(* Logix 5000 project; controller FV vendor 1 type 14 code 217 rev 31.11; software revision 31.00; part 7 of 63 *)
(* tags used below, declared in another part *)
   CWD : CHECKWORD_FLAGS;
   Dummy : BOOL;
   FR_B240 : INT[255];   // DEBOUNCE Debounce Flags
   fr_chk_temp : DINT;
   FR_copy_how_many : DINT;
   FR_data_file_value_to_move : DINT;
   FR_from_data_file : DINT;
   FR_from_data_offset : DINT;
   FR_FV26_HLP01 : PlantItem;   // FV26_HLP01
   FR_FV26_LLP01 : PlantItem;   // FV26_LLP01
   FR_FV27_HLP01 : PlantItem;   // FV27_HLP01
   FR_FV27_LLP01 : PlantItem;   // FV27_LLP01
   FR_FV28_HLP01 : PlantItem;   // FV28_HLP01
   FR_FV28_LLP01 : PlantItem;   // FV28_LLP01
   FR_FV29_HLP01 : PlantItem;   // FV29_HLP01
   FR_FV29_LLP01 : PlantItem;   // FV29_LLP01
   FR_FV30_HLP01 : PlantItem;   // FV30_HLP01
   FR_FV30_LLP01 : PlantItem;   // FV30_LLP01
   FR_FV31_HLP01 : PlantItem;   // FV31_HLP01
   FR_N10 : INT[265];   // FV_AGING Comms to FV Aging PL C
   FR_N100 : INT[265];   // FV FILLING
   FR_N110 : INT[265];   // GREEN BEER Green Beer Main
   FR_N120 : INT[265];   // YEAST CROP Yeast Cropping Main
   FR_N13 : INT[265];   // MV_ROUTE Comms to MV Routing PLC
   FR_N130 : INT[265];   // FILTRATE Filtrate Return
   FR_N14 : INT[265];   // MVFV CIP Comms to MVFV CIP Un it PLC
   FR_N140 : INT[265];   // CIP
   FR_N142 : INT[265];   // CIP
   FR_N143 : INT[265];   // CIP
   FR_N150 : INT[265];   // Original N File From SLC, No Description Available
   FR_N160 : INT[265];   // VESSEL Vessel Working Direc tory
   FR_N170 : INT[265];   // Original N File From SLC, No Description Available
   FR_N180 : INT[265];   // Original N File From SLC, No Description Available
   FR_N198 : INT[265];   // Original N File From SLC, No Description Available
   FR_N20 : INT[265];   // GENERAL General Purpose Setp oints
   FR_N200 : INT[265];   // ANALOG_IN Analog Inputs
   FR_N201 : INT[265];   // Original N File From SLC, No Description Available
   FR_N207 : INT[265];   // Original N File From SLC, No Description Available
   FR_N21 : INT[265];   // CHASE_V FV Filling Beer Chas e Volumes
   FR_N210 : INT[265];   // ANALOG_OUT Analog Outputs
   FR_N220 : INT[265];   // CHECKLIST Checklist Loop Contr ollers
   FR_N225 : INT[265];   // Original N File From SLC, No Description Available
   FR_N226 : INT[265];   // Original N File From SLC, No Description Available
   FR_N245 : INT[265];   // CHECKWORD Checkword Loop Contr ol
   FR_N252 : INT[265];   // OUTPUT_PTR Checkword Pointers t o output flags in B2 50
   FR_N253 : INT[265];   // EN_POINT Pointers to energise d input flags in B25 1
   FR_N254 : INT[265];   // DEN_POINT Pointers to deenergi sed input flags in B 251
   FR_N255 : INT[265];   // CHECKWORDS
   FR_N26 : INT[265];   // FV26
   FR_N27 : INT[265];   // FV27
   FR_N28 : INT[265];   // FV28
   FR_N29 : INT[265];   // FV29
   FR_N30 : INT[265];   // FV30
   FR_N31 : INT[265];   // FV31
   FR_N36 : INT[265];   // Original N File From SLC, No Description Available
   FR_N37 : INT[265];   // Original N File From SLC, No Description Available
   FR_N46 : INT[265];   // Original N File From SLC, No Description Available
   FR_N47 : INT[265];   // Original N File From SLC, No Description Available
   FR_N7 : INT[265];   // INTEGER
   FR_N99 : INT[265];   // COMMENT Comment Lines
   FR_T242 : TIMER[255];   // DEBOUNCE
   FR_T243 : TIMER[255];   // DEBOUNCE
   FR_to_data_file : DINT;
   FR_to_data_offset : DINT;
(* FR_Common, continued *)

ROUTINE FR_CHECK_LIST_220   (* ladder *)
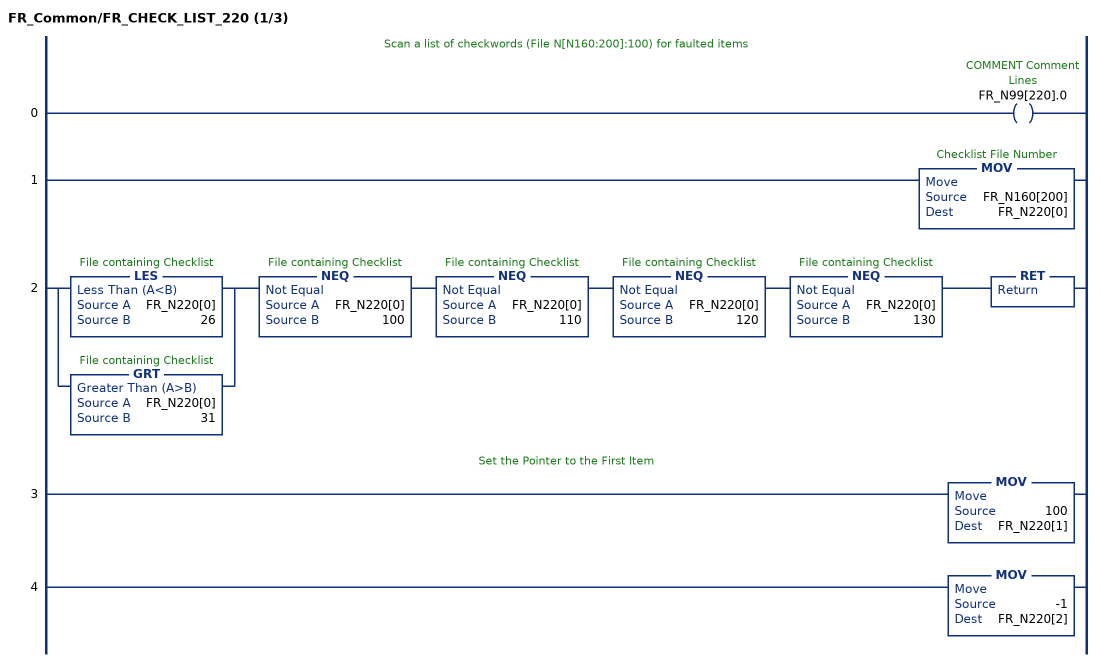
   // Scan a list of checkwords (File N[N160:200]:100) for faulted items
   0: OTE(FR_N99[220].0);
   1: MOV(FR_N160[200],FR_N220[0]);
   2: [LES(FR_N220[0],26) ,GRT(FR_N220[0],31) ]NEQ(FR_N220[0],100)NEQ(FR_N220[0],110)NEQ(FR_N220[0],120)NEQ(FR_N220[0],130)RET();
   // Set the Pointer to the First Item
   3: MOV(100,FR_N220[1]);
   4: MOV(-1,FR_N220[2]);
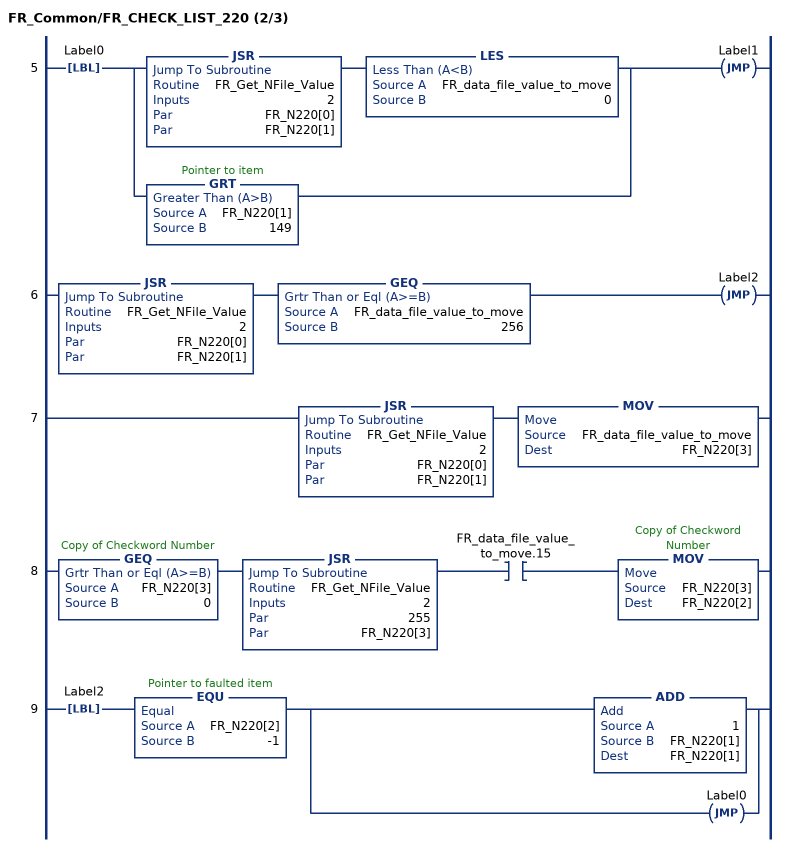
   5: LBL(Label0)[JSR(FR_Get_NFile_Value,2,FR_N220[0],FR_N220[1]) LES(FR_data_file_value_to_move,0) ,GRT(FR_N220[1],149) ]JMP(Label1);
   6: JSR(FR_Get_NFile_Value,2,FR_N220[0],FR_N220[1])GEQ(FR_data_file_value_to_move,256)JMP(Label2);
   7: JSR(FR_Get_NFile_Value,2,FR_N220[0],FR_N220[1])MOV(FR_data_file_value_to_move,FR_N220[3]);
   8: GEQ(FR_N220[3],0)JSR(FR_Get_NFile_Value,2,255,FR_N220[3])XIC(FR_data_file_value_to_move.15)MOV(FR_N220[3],FR_N220[2]);
   9: LBL(Label2)EQU(FR_N220[2],-1)[ADD(1,FR_N220[1],FR_N220[1]) ,JMP(Label0) ];
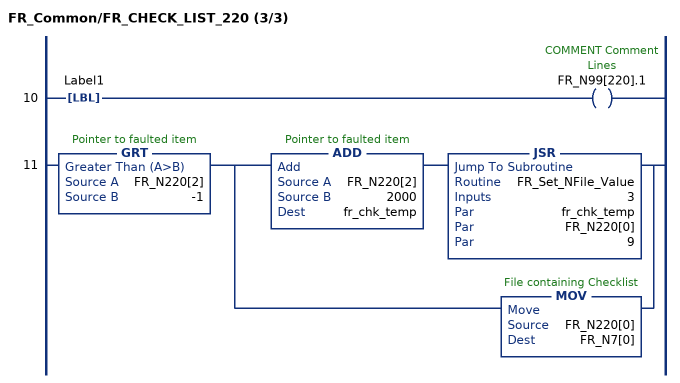
   10: LBL(Label1)OTE(FR_N99[220].1);
   11: GRT(FR_N220[2],-1)[ADD(FR_N220[2],2000,fr_chk_temp) JSR(FR_Set_NFile_Value,3,fr_chk_temp,FR_N220[0],9) ,MOV(FR_N220[0],FR_N7[0]) ];
END_ROUTINE

ROUTINE FR_CHECKRESET_221   (* ladder *)
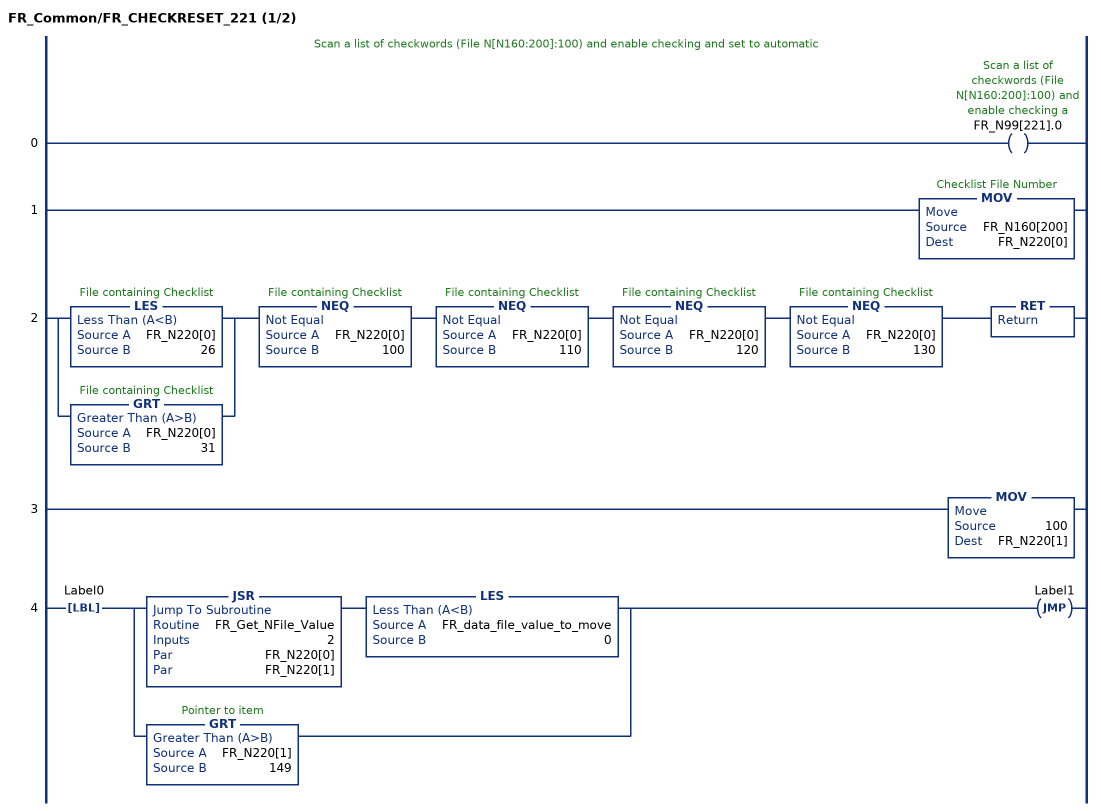
   // Scan a list of checkwords (File N[N160:200]:100) and enable checking and set to automatic
   0: OTE(FR_N99[221].0);
   1: MOV(FR_N160[200],FR_N220[0]);
   2: [LES(FR_N220[0],26) ,GRT(FR_N220[0],31) ]NEQ(FR_N220[0],100)NEQ(FR_N220[0],110)NEQ(FR_N220[0],120)NEQ(FR_N220[0],130)RET();
   3: MOV(100,FR_N220[1]);
   4: LBL(Label0)[JSR(FR_Get_NFile_Value,2,FR_N220[0],FR_N220[1]) LES(FR_data_file_value_to_move,0) ,GRT(FR_N220[1],149) ]JMP(Label1);
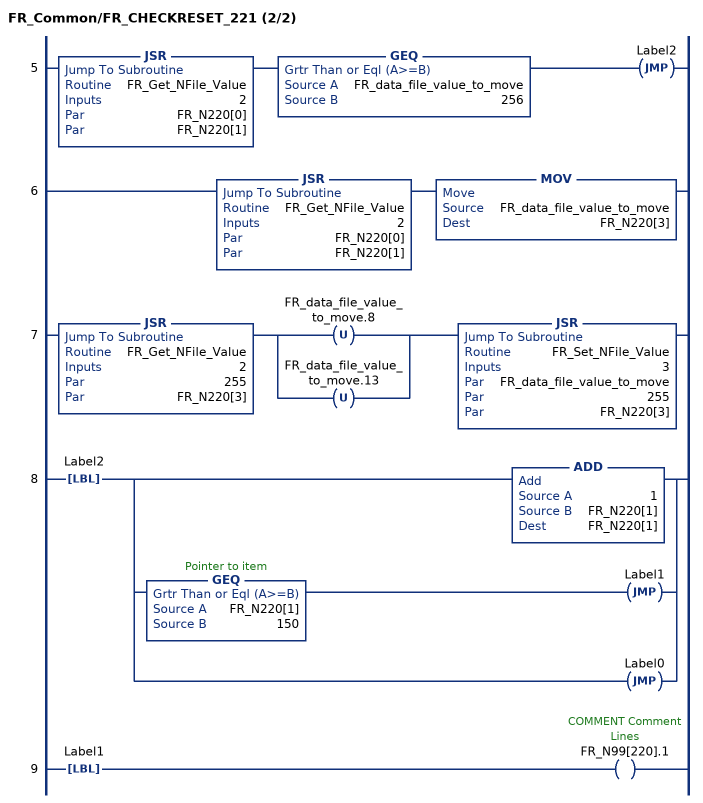
   5: JSR(FR_Get_NFile_Value,2,FR_N220[0],FR_N220[1])GEQ(FR_data_file_value_to_move,256)JMP(Label2);
   6: JSR(FR_Get_NFile_Value,2,FR_N220[0],FR_N220[1])MOV(FR_data_file_value_to_move,FR_N220[3]);
   7: JSR(FR_Get_NFile_Value,2,255,FR_N220[3])[OTU(FR_data_file_value_to_move.8) ,OTU(FR_data_file_value_to_move.13) ]JSR(FR_Set_NFile_Value,3,FR_data_file_value_to_move,255,FR_N220[3]);
   8: LBL(Label2)[ADD(1,FR_N220[1],FR_N220[1]) ,GEQ(FR_N220[1],150) JMP(Label1) ,JMP(Label0) ];
   9: LBL(Label1)OTE(FR_N99[220].1);
END_ROUTINE

ROUTINE FR_Copy_NFile_Block   (* ladder *)
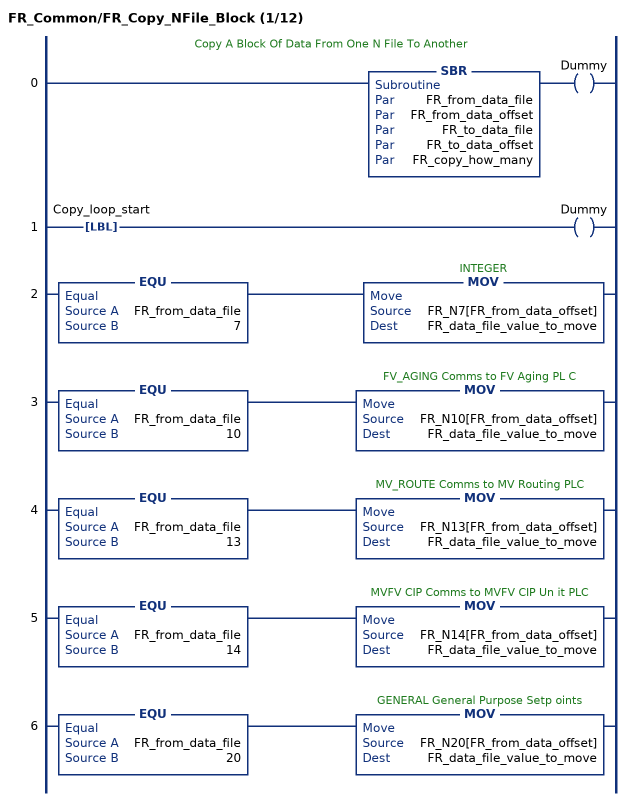
   // Copy A Block Of Data From One N File To Another
   0: SBR(FR_from_data_file,FR_from_data_offset,FR_to_data_file,FR_to_data_offset,FR_copy_how_many)OTE(Dummy);
   1: LBL(Copy_loop_start)OTE(Dummy);
   2: EQU(FR_from_data_file,7)MOV(FR_N7[FR_from_data_offset],FR_data_file_value_to_move);
   3: EQU(FR_from_data_file,10)MOV(FR_N10[FR_from_data_offset],FR_data_file_value_to_move);
   4: EQU(FR_from_data_file,13)MOV(FR_N13[FR_from_data_offset],FR_data_file_value_to_move);
   5: EQU(FR_from_data_file,14)MOV(FR_N14[FR_from_data_offset],FR_data_file_value_to_move);
   6: EQU(FR_from_data_file,20)MOV(FR_N20[FR_from_data_offset],FR_data_file_value_to_move);
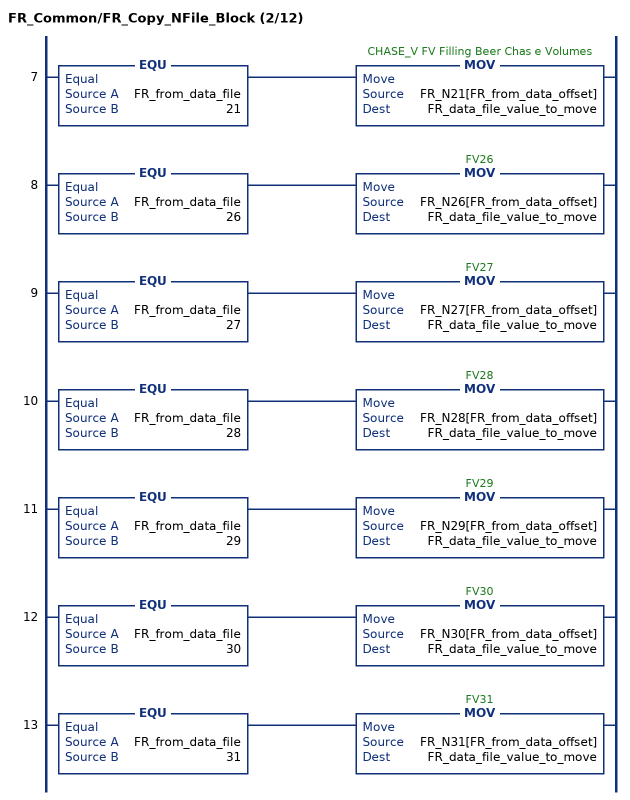
   7: EQU(FR_from_data_file,21)MOV(FR_N21[FR_from_data_offset],FR_data_file_value_to_move);
   8: EQU(FR_from_data_file,26)MOV(FR_N26[FR_from_data_offset],FR_data_file_value_to_move);
   9: EQU(FR_from_data_file,27)MOV(FR_N27[FR_from_data_offset],FR_data_file_value_to_move);
   10: EQU(FR_from_data_file,28)MOV(FR_N28[FR_from_data_offset],FR_data_file_value_to_move);
   11: EQU(FR_from_data_file,29)MOV(FR_N29[FR_from_data_offset],FR_data_file_value_to_move);
   12: EQU(FR_from_data_file,30)MOV(FR_N30[FR_from_data_offset],FR_data_file_value_to_move);
   13: EQU(FR_from_data_file,31)MOV(FR_N31[FR_from_data_offset],FR_data_file_value_to_move);
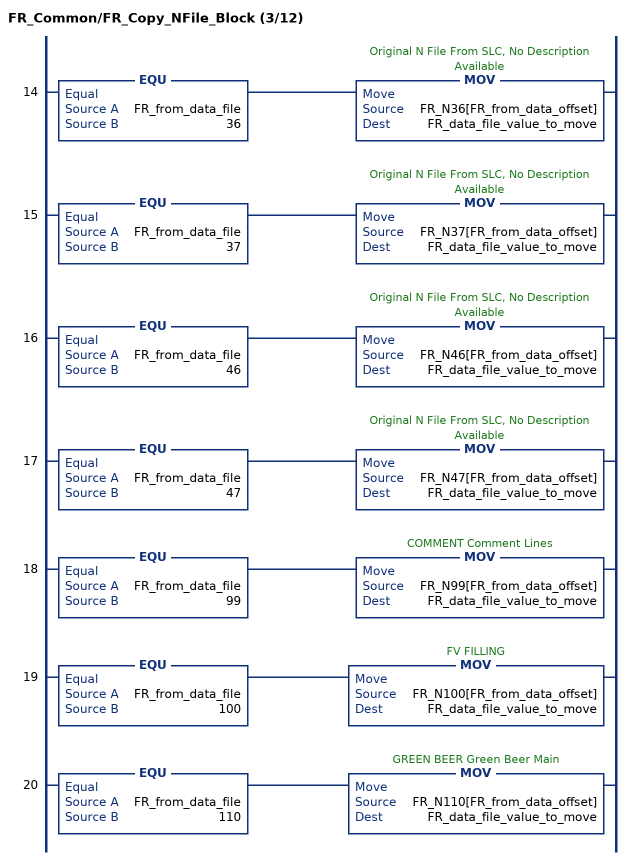
   14: EQU(FR_from_data_file,36)MOV(FR_N36[FR_from_data_offset],FR_data_file_value_to_move);
   15: EQU(FR_from_data_file,37)MOV(FR_N37[FR_from_data_offset],FR_data_file_value_to_move);
   16: EQU(FR_from_data_file,46)MOV(FR_N46[FR_from_data_offset],FR_data_file_value_to_move);
   17: EQU(FR_from_data_file,47)MOV(FR_N47[FR_from_data_offset],FR_data_file_value_to_move);
   18: EQU(FR_from_data_file,99)MOV(FR_N99[FR_from_data_offset],FR_data_file_value_to_move);
   19: EQU(FR_from_data_file,100)MOV(FR_N100[FR_from_data_offset],FR_data_file_value_to_move);
   20: EQU(FR_from_data_file,110)MOV(FR_N110[FR_from_data_offset],FR_data_file_value_to_move);
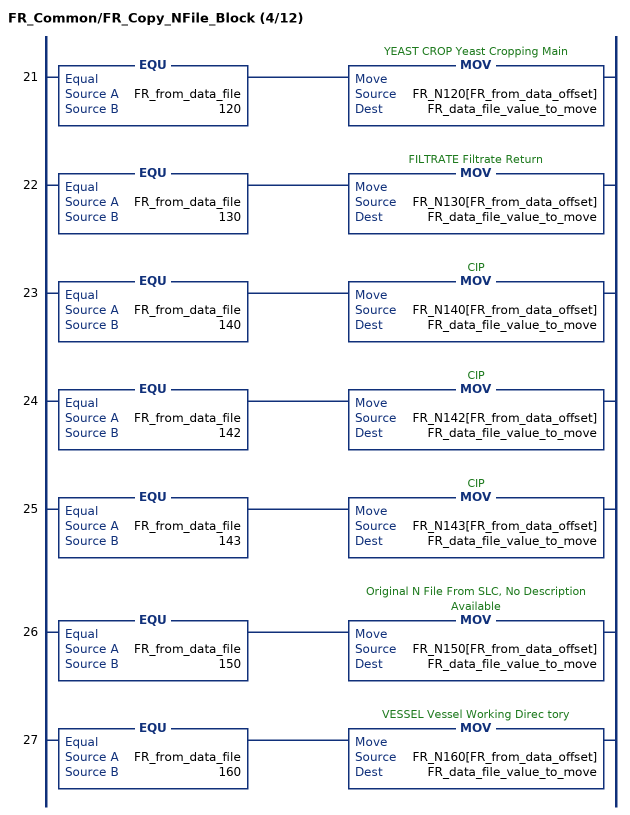
   21: EQU(FR_from_data_file,120)MOV(FR_N120[FR_from_data_offset],FR_data_file_value_to_move);
   22: EQU(FR_from_data_file,130)MOV(FR_N130[FR_from_data_offset],FR_data_file_value_to_move);
   23: EQU(FR_from_data_file,140)MOV(FR_N140[FR_from_data_offset],FR_data_file_value_to_move);
   24: EQU(FR_from_data_file,142)MOV(FR_N142[FR_from_data_offset],FR_data_file_value_to_move);
   25: EQU(FR_from_data_file,143)MOV(FR_N143[FR_from_data_offset],FR_data_file_value_to_move);
   26: EQU(FR_from_data_file,150)MOV(FR_N150[FR_from_data_offset],FR_data_file_value_to_move);
   27: EQU(FR_from_data_file,160)MOV(FR_N160[FR_from_data_offset],FR_data_file_value_to_move);
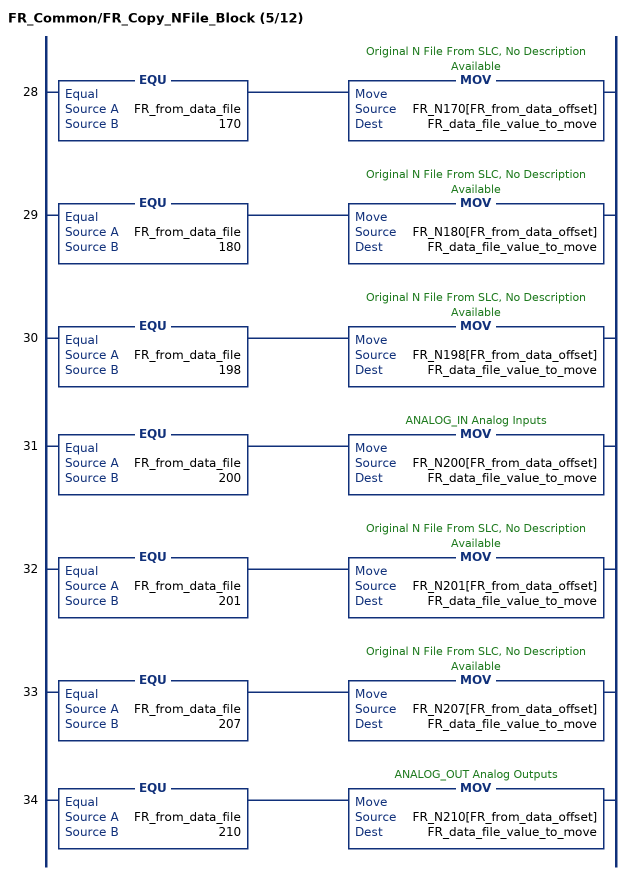
   28: EQU(FR_from_data_file,170)MOV(FR_N170[FR_from_data_offset],FR_data_file_value_to_move);
   29: EQU(FR_from_data_file,180)MOV(FR_N180[FR_from_data_offset],FR_data_file_value_to_move);
   30: EQU(FR_from_data_file,198)MOV(FR_N198[FR_from_data_offset],FR_data_file_value_to_move);
   31: EQU(FR_from_data_file,200)MOV(FR_N200[FR_from_data_offset],FR_data_file_value_to_move);
   32: EQU(FR_from_data_file,201)MOV(FR_N201[FR_from_data_offset],FR_data_file_value_to_move);
   33: EQU(FR_from_data_file,207)MOV(FR_N207[FR_from_data_offset],FR_data_file_value_to_move);
   34: EQU(FR_from_data_file,210)MOV(FR_N210[FR_from_data_offset],FR_data_file_value_to_move);
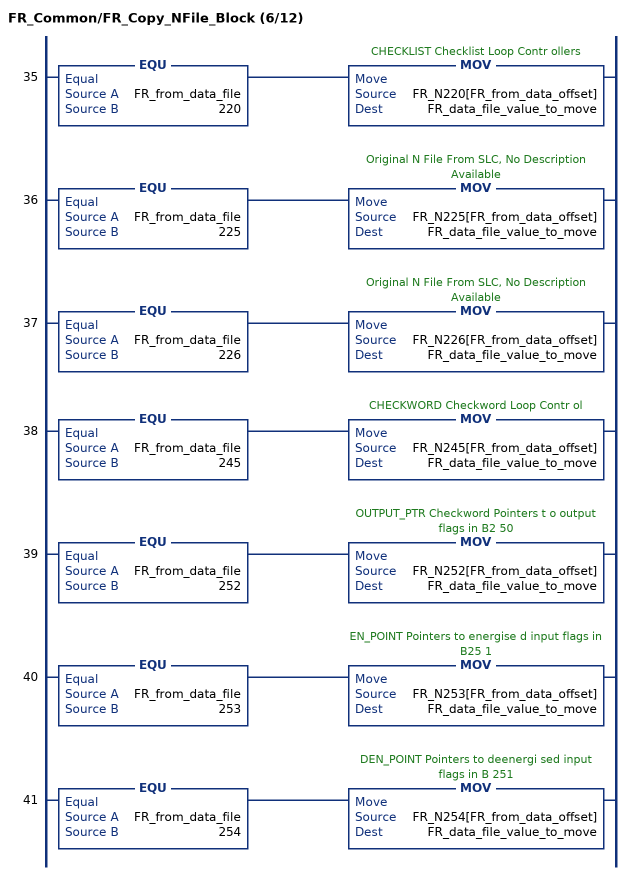
   35: EQU(FR_from_data_file,220)MOV(FR_N220[FR_from_data_offset],FR_data_file_value_to_move);
   36: EQU(FR_from_data_file,225)MOV(FR_N225[FR_from_data_offset],FR_data_file_value_to_move);
   37: EQU(FR_from_data_file,226)MOV(FR_N226[FR_from_data_offset],FR_data_file_value_to_move);
   38: EQU(FR_from_data_file,245)MOV(FR_N245[FR_from_data_offset],FR_data_file_value_to_move);
   39: EQU(FR_from_data_file,252)MOV(FR_N252[FR_from_data_offset],FR_data_file_value_to_move);
   40: EQU(FR_from_data_file,253)MOV(FR_N253[FR_from_data_offset],FR_data_file_value_to_move);
   41: EQU(FR_from_data_file,254)MOV(FR_N254[FR_from_data_offset],FR_data_file_value_to_move);
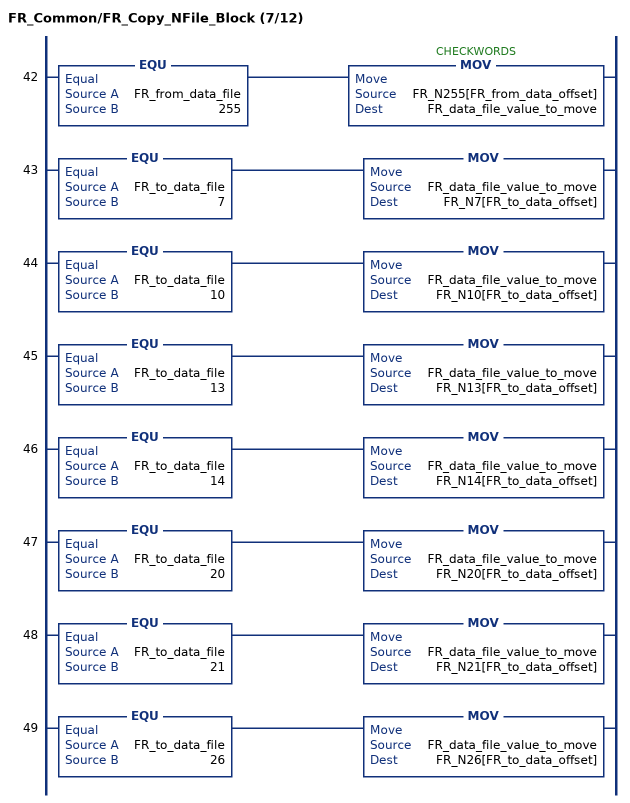
   42: EQU(FR_from_data_file,255)MOV(FR_N255[FR_from_data_offset],FR_data_file_value_to_move);
   43: EQU(FR_to_data_file,7)MOV(FR_data_file_value_to_move,FR_N7[FR_to_data_offset]);
   44: EQU(FR_to_data_file,10)MOV(FR_data_file_value_to_move,FR_N10[FR_to_data_offset]);
   45: EQU(FR_to_data_file,13)MOV(FR_data_file_value_to_move,FR_N13[FR_to_data_offset]);
   46: EQU(FR_to_data_file,14)MOV(FR_data_file_value_to_move,FR_N14[FR_to_data_offset]);
   47: EQU(FR_to_data_file,20)MOV(FR_data_file_value_to_move,FR_N20[FR_to_data_offset]);
   48: EQU(FR_to_data_file,21)MOV(FR_data_file_value_to_move,FR_N21[FR_to_data_offset]);
   49: EQU(FR_to_data_file,26)MOV(FR_data_file_value_to_move,FR_N26[FR_to_data_offset]);
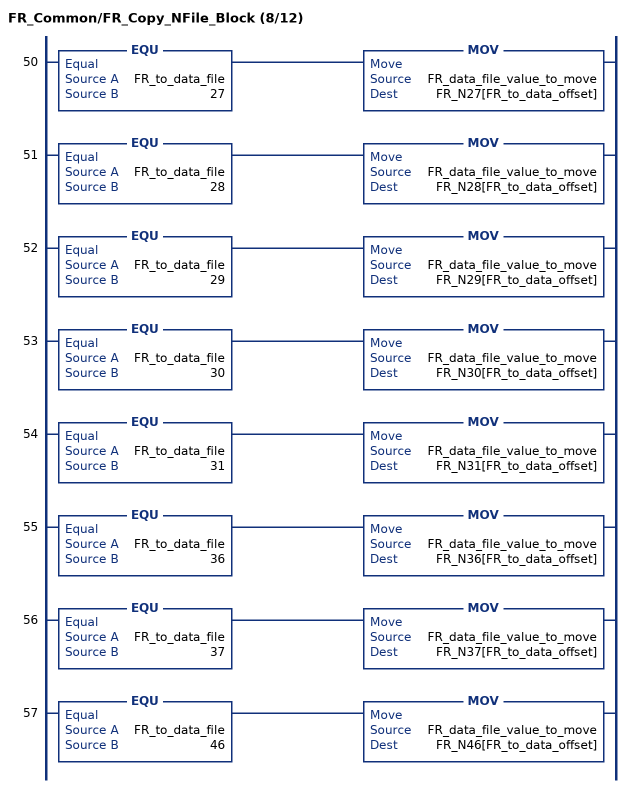
   50: EQU(FR_to_data_file,27)MOV(FR_data_file_value_to_move,FR_N27[FR_to_data_offset]);
   51: EQU(FR_to_data_file,28)MOV(FR_data_file_value_to_move,FR_N28[FR_to_data_offset]);
   52: EQU(FR_to_data_file,29)MOV(FR_data_file_value_to_move,FR_N29[FR_to_data_offset]);
   53: EQU(FR_to_data_file,30)MOV(FR_data_file_value_to_move,FR_N30[FR_to_data_offset]);
   54: EQU(FR_to_data_file,31)MOV(FR_data_file_value_to_move,FR_N31[FR_to_data_offset]);
   55: EQU(FR_to_data_file,36)MOV(FR_data_file_value_to_move,FR_N36[FR_to_data_offset]);
   56: EQU(FR_to_data_file,37)MOV(FR_data_file_value_to_move,FR_N37[FR_to_data_offset]);
   57: EQU(FR_to_data_file,46)MOV(FR_data_file_value_to_move,FR_N46[FR_to_data_offset]);
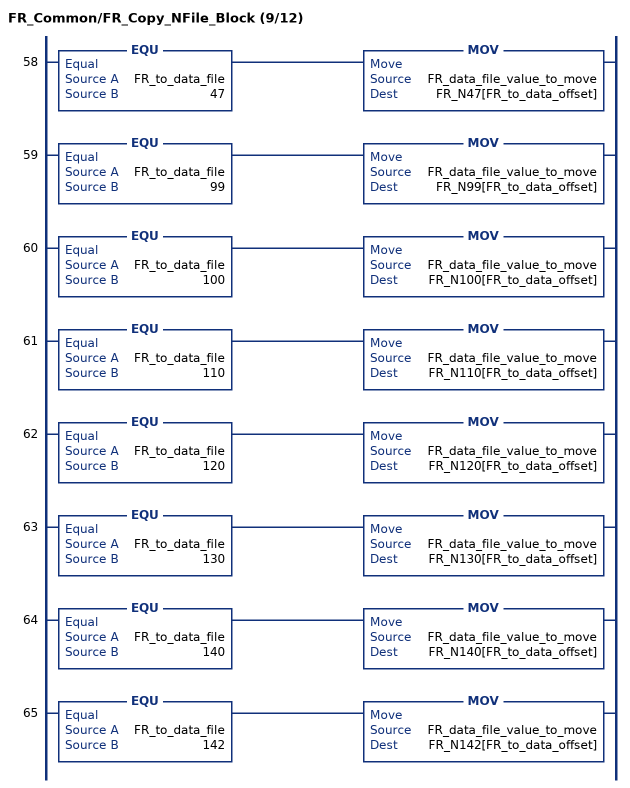
   58: EQU(FR_to_data_file,47)MOV(FR_data_file_value_to_move,FR_N47[FR_to_data_offset]);
   59: EQU(FR_to_data_file,99)MOV(FR_data_file_value_to_move,FR_N99[FR_to_data_offset]);
   60: EQU(FR_to_data_file,100)MOV(FR_data_file_value_to_move,FR_N100[FR_to_data_offset]);
   61: EQU(FR_to_data_file,110)MOV(FR_data_file_value_to_move,FR_N110[FR_to_data_offset]);
   62: EQU(FR_to_data_file,120)MOV(FR_data_file_value_to_move,FR_N120[FR_to_data_offset]);
   63: EQU(FR_to_data_file,130)MOV(FR_data_file_value_to_move,FR_N130[FR_to_data_offset]);
   64: EQU(FR_to_data_file,140)MOV(FR_data_file_value_to_move,FR_N140[FR_to_data_offset]);
   65: EQU(FR_to_data_file,142)MOV(FR_data_file_value_to_move,FR_N142[FR_to_data_offset]);
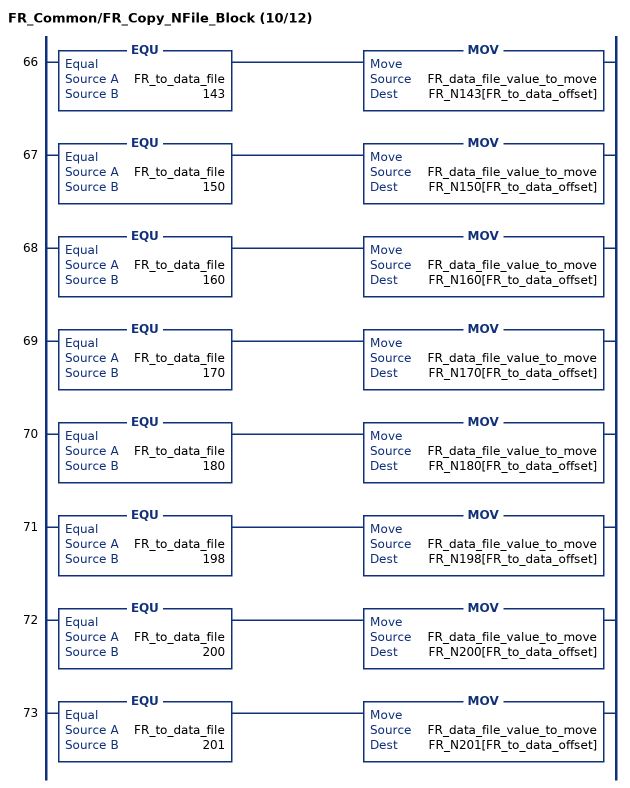
   66: EQU(FR_to_data_file,143)MOV(FR_data_file_value_to_move,FR_N143[FR_to_data_offset]);
   67: EQU(FR_to_data_file,150)MOV(FR_data_file_value_to_move,FR_N150[FR_to_data_offset]);
   68: EQU(FR_to_data_file,160)MOV(FR_data_file_value_to_move,FR_N160[FR_to_data_offset]);
   69: EQU(FR_to_data_file,170)MOV(FR_data_file_value_to_move,FR_N170[FR_to_data_offset]);
   70: EQU(FR_to_data_file,180)MOV(FR_data_file_value_to_move,FR_N180[FR_to_data_offset]);
   71: EQU(FR_to_data_file,198)MOV(FR_data_file_value_to_move,FR_N198[FR_to_data_offset]);
   72: EQU(FR_to_data_file,200)MOV(FR_data_file_value_to_move,FR_N200[FR_to_data_offset]);
   73: EQU(FR_to_data_file,201)MOV(FR_data_file_value_to_move,FR_N201[FR_to_data_offset]);
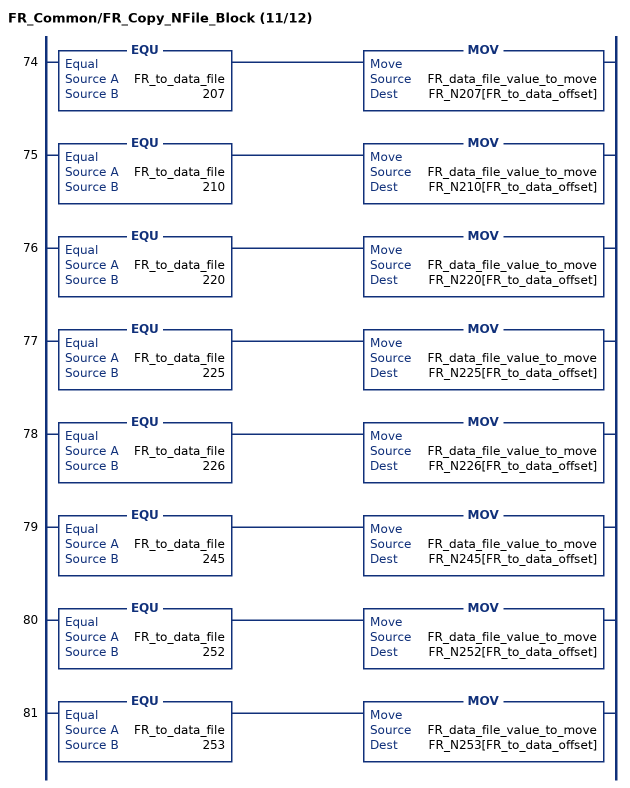
   74: EQU(FR_to_data_file,207)MOV(FR_data_file_value_to_move,FR_N207[FR_to_data_offset]);
   75: EQU(FR_to_data_file,210)MOV(FR_data_file_value_to_move,FR_N210[FR_to_data_offset]);
   76: EQU(FR_to_data_file,220)MOV(FR_data_file_value_to_move,FR_N220[FR_to_data_offset]);
   77: EQU(FR_to_data_file,225)MOV(FR_data_file_value_to_move,FR_N225[FR_to_data_offset]);
   78: EQU(FR_to_data_file,226)MOV(FR_data_file_value_to_move,FR_N226[FR_to_data_offset]);
   79: EQU(FR_to_data_file,245)MOV(FR_data_file_value_to_move,FR_N245[FR_to_data_offset]);
   80: EQU(FR_to_data_file,252)MOV(FR_data_file_value_to_move,FR_N252[FR_to_data_offset]);
   81: EQU(FR_to_data_file,253)MOV(FR_data_file_value_to_move,FR_N253[FR_to_data_offset]);
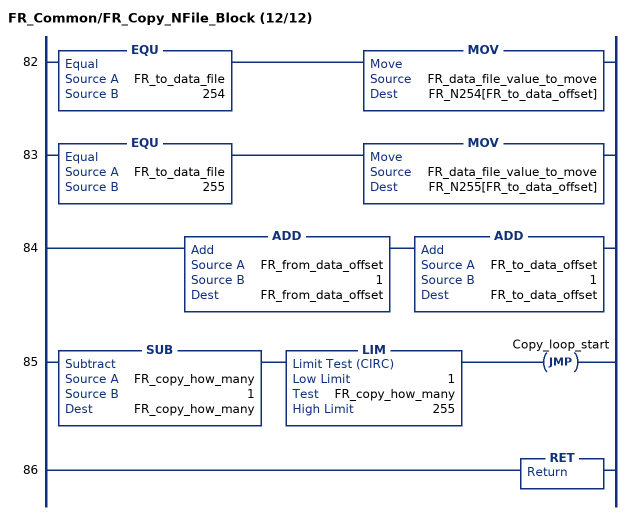
   82: EQU(FR_to_data_file,254)MOV(FR_data_file_value_to_move,FR_N254[FR_to_data_offset]);
   83: EQU(FR_to_data_file,255)MOV(FR_data_file_value_to_move,FR_N255[FR_to_data_offset]);
   84: ADD(FR_from_data_offset,1,FR_from_data_offset)ADD(FR_to_data_offset,1,FR_to_data_offset);
   85: SUB(FR_copy_how_many,1,FR_copy_how_many)LIM(1,FR_copy_how_many,255)JMP(Copy_loop_start);
   86: RET();
END_ROUTINE

ROUTINE FR_DEBOUNCE_240   (* ladder *)
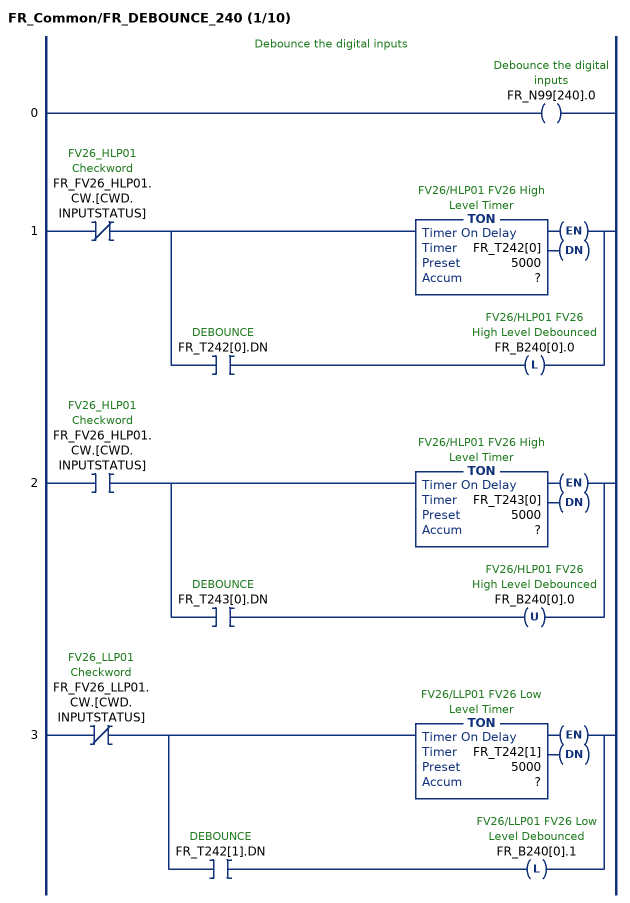
   // Debounce the digital inputs
   0: OTE(FR_N99[240].0);
   1: XIO(FR_FV26_HLP01.CW.[CWD.INPUTSTATUS])[TON(FR_T242[0],?,?) ,XIC(FR_T242[0].DN) OTL(FR_B240[0].0) ];
   2: XIC(FR_FV26_HLP01.CW.[CWD.INPUTSTATUS])[TON(FR_T243[0],?,?) ,XIC(FR_T243[0].DN) OTU(FR_B240[0].0) ];
   3: XIO(FR_FV26_LLP01.CW.[CWD.INPUTSTATUS])[TON(FR_T242[1],?,?) ,XIC(FR_T242[1].DN) OTL(FR_B240[0].1) ];
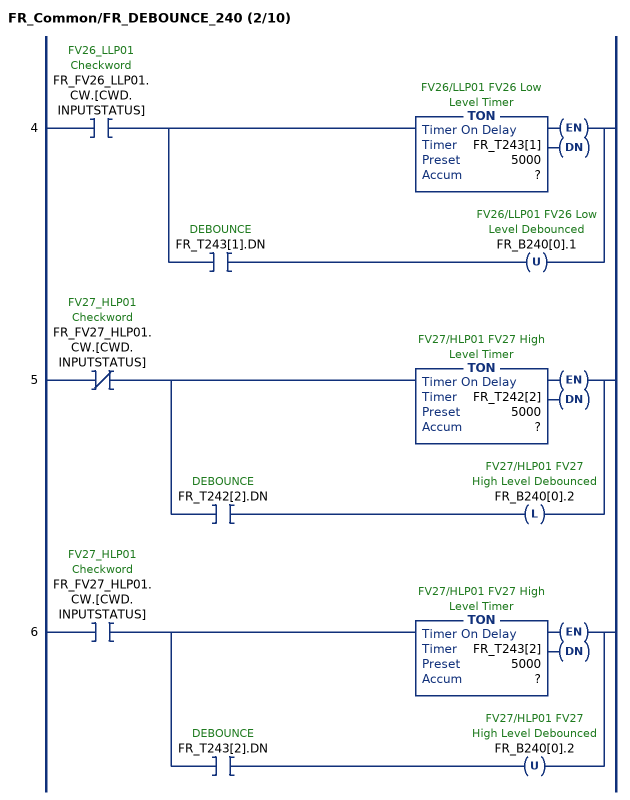
   4: XIC(FR_FV26_LLP01.CW.[CWD.INPUTSTATUS])[TON(FR_T243[1],?,?) ,XIC(FR_T243[1].DN) OTU(FR_B240[0].1) ];
   5: XIO(FR_FV27_HLP01.CW.[CWD.INPUTSTATUS])[TON(FR_T242[2],?,?) ,XIC(FR_T242[2].DN) OTL(FR_B240[0].2) ];
   6: XIC(FR_FV27_HLP01.CW.[CWD.INPUTSTATUS])[TON(FR_T243[2],?,?) ,XIC(FR_T243[2].DN) OTU(FR_B240[0].2) ];
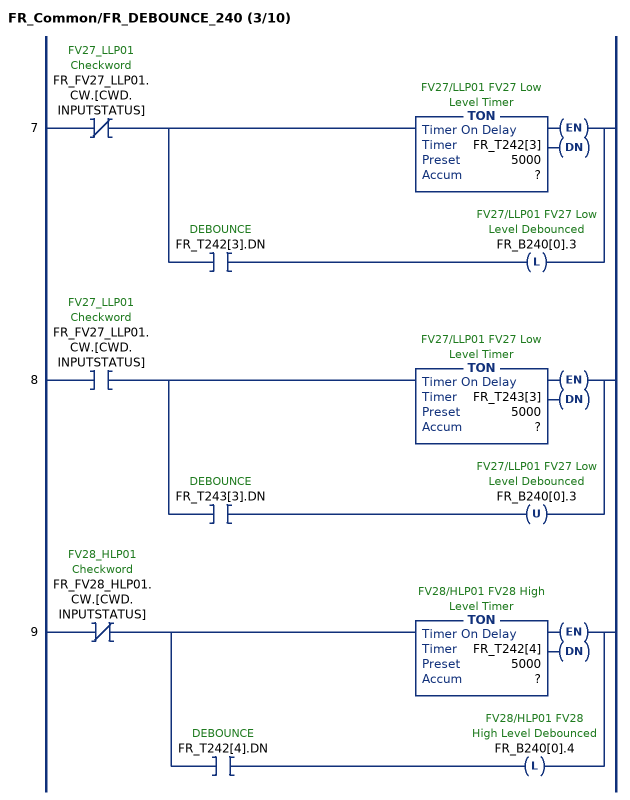
   7: XIO(FR_FV27_LLP01.CW.[CWD.INPUTSTATUS])[TON(FR_T242[3],?,?) ,XIC(FR_T242[3].DN) OTL(FR_B240[0].3) ];
   8: XIC(FR_FV27_LLP01.CW.[CWD.INPUTSTATUS])[TON(FR_T243[3],?,?) ,XIC(FR_T243[3].DN) OTU(FR_B240[0].3) ];
   9: XIO(FR_FV28_HLP01.CW.[CWD.INPUTSTATUS])[TON(FR_T242[4],?,?) ,XIC(FR_T242[4].DN) OTL(FR_B240[0].4) ];
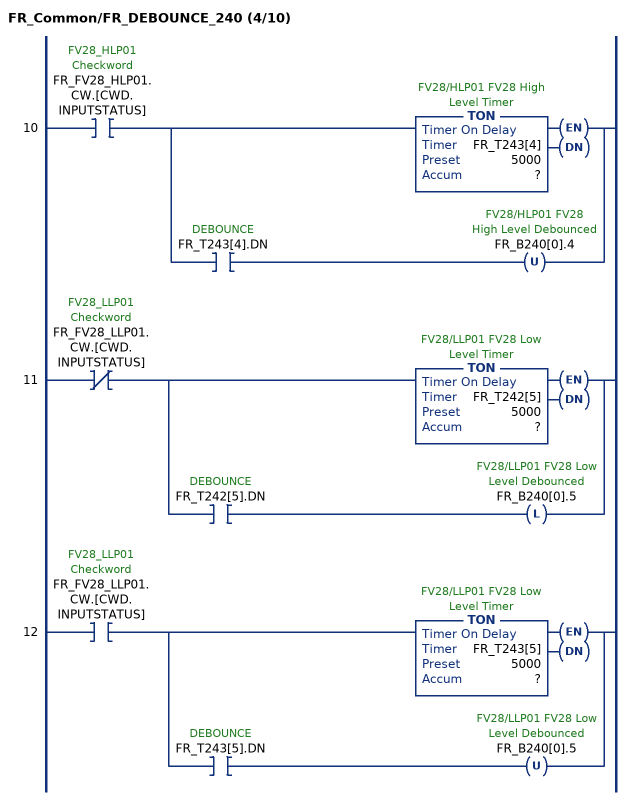
   10: XIC(FR_FV28_HLP01.CW.[CWD.INPUTSTATUS])[TON(FR_T243[4],?,?) ,XIC(FR_T243[4].DN) OTU(FR_B240[0].4) ];
   11: XIO(FR_FV28_LLP01.CW.[CWD.INPUTSTATUS])[TON(FR_T242[5],?,?) ,XIC(FR_T242[5].DN) OTL(FR_B240[0].5) ];
   12: XIC(FR_FV28_LLP01.CW.[CWD.INPUTSTATUS])[TON(FR_T243[5],?,?) ,XIC(FR_T243[5].DN) OTU(FR_B240[0].5) ];
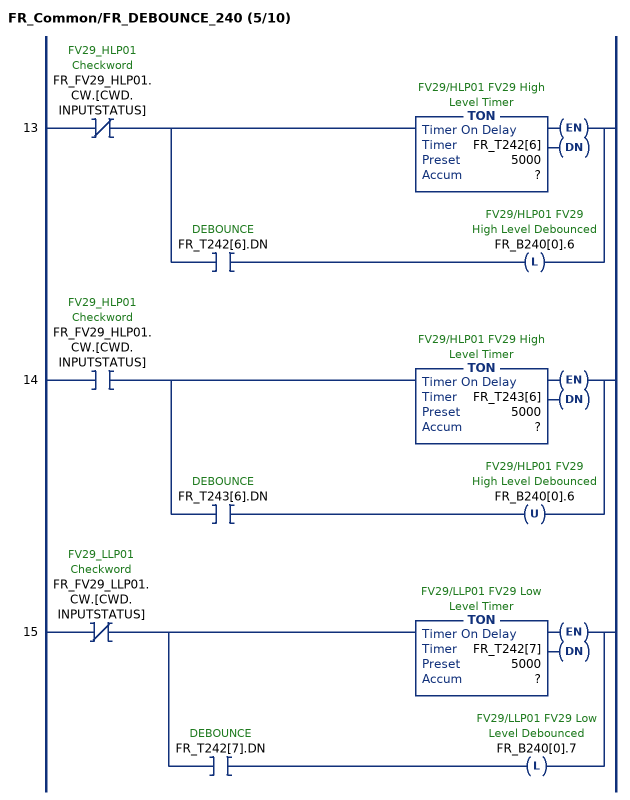
   13: XIO(FR_FV29_HLP01.CW.[CWD.INPUTSTATUS])[TON(FR_T242[6],?,?) ,XIC(FR_T242[6].DN) OTL(FR_B240[0].6) ];
   14: XIC(FR_FV29_HLP01.CW.[CWD.INPUTSTATUS])[TON(FR_T243[6],?,?) ,XIC(FR_T243[6].DN) OTU(FR_B240[0].6) ];
   15: XIO(FR_FV29_LLP01.CW.[CWD.INPUTSTATUS])[TON(FR_T242[7],?,?) ,XIC(FR_T242[7].DN) OTL(FR_B240[0].7) ];
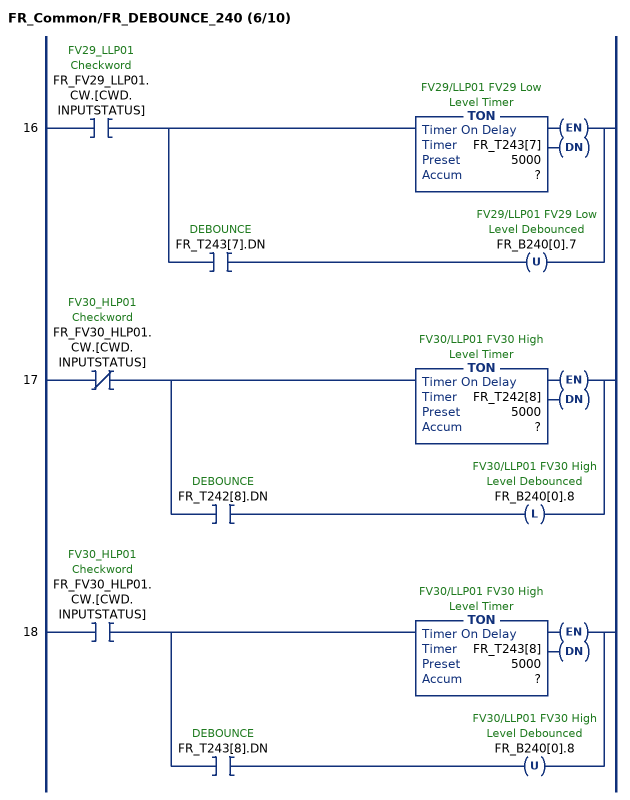
   16: XIC(FR_FV29_LLP01.CW.[CWD.INPUTSTATUS])[TON(FR_T243[7],?,?) ,XIC(FR_T243[7].DN) OTU(FR_B240[0].7) ];
   17: XIO(FR_FV30_HLP01.CW.[CWD.INPUTSTATUS])[TON(FR_T242[8],?,?) ,XIC(FR_T242[8].DN) OTL(FR_B240[0].8) ];
   18: XIC(FR_FV30_HLP01.CW.[CWD.INPUTSTATUS])[TON(FR_T243[8],?,?) ,XIC(FR_T243[8].DN) OTU(FR_B240[0].8) ];
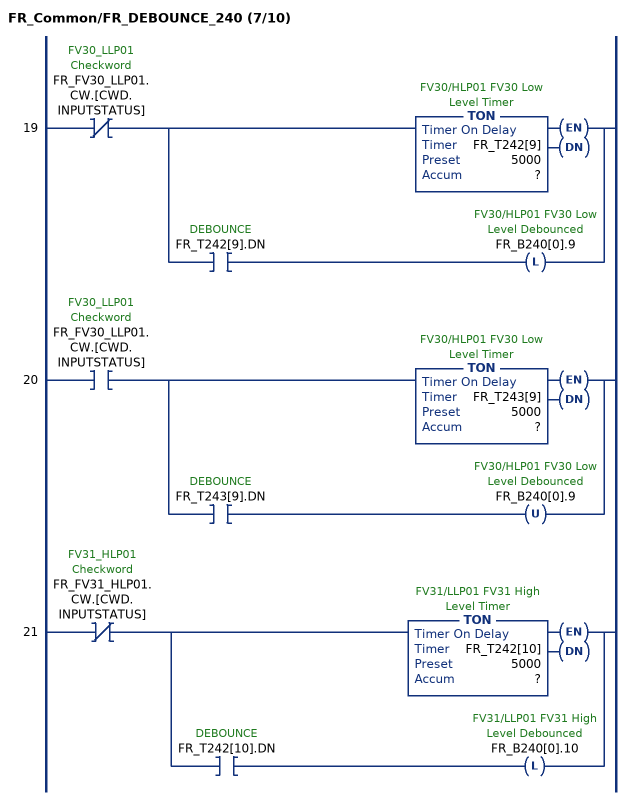
   19: XIO(FR_FV30_LLP01.CW.[CWD.INPUTSTATUS])[TON(FR_T242[9],?,?) ,XIC(FR_T242[9].DN) OTL(FR_B240[0].9) ];
   20: XIC(FR_FV30_LLP01.CW.[CWD.INPUTSTATUS])[TON(FR_T243[9],?,?) ,XIC(FR_T243[9].DN) OTU(FR_B240[0].9) ];
   21: XIO(FR_FV31_HLP01.CW.[CWD.INPUTSTATUS])[TON(FR_T242[10],?,?) ,XIC(FR_T242[10].DN) OTL(FR_B240[0].10) ];
